// TIA Portal project "Respirator2020_V16" (V16)

(* hardware
DEVICE "S7-1200 station_1"  S7-1200 Station
   slot 0: "Rack_0"  S7-1200 Rack  Rack  V1.0
   slot 1: "PLC_1"  CPU 1215C DC/DC/DC  6ES7 215-1AG40-0XB0  V4.2
DEVICE "HMI_1"  TP700 Comfort
   slot 0: "HMI_1"  TP700 Comfort  6AV2 124-0GC01-0AX0  15.1.0.0
   slot 1: "HMI_RT_1"  TP700 Comfort  6AV2 124-0GC01-0AX0  15.1.0.0
   slot 5: "HMI_1.IE_CP_1"  PROFINET Interface  15.0.1.0
      slot 1: "Interfaz PROFINET_1"  PROFINET Interface
         slot 1: "Port_1"  Port
         slot 2: "Port_2"  Port
   slot 7: "HMI_1.MPI/DP_CP_1"  MPI/DP Interface  15.0.1.0
*)

// ===== PLC "PLC_1"  CPU 1215C DC/DC/DC =====

VAR_GLOBAL   // PLC tag table "Tabla de variables estándar"
   "System_Byte" AT %MB1 : Byte;
   "FirstScan" AT %M1.0 : Bool;
   "DiagStatusUpdate" AT %M1.1 : Bool;
   "AlwaysTRUE" AT %M1.2 : Bool;
   "AlwaysFALSE" AT %M1.3 : Bool;
   "Clock_Byte" AT %MB0 : Byte;
   "Clock_10Hz" AT %M0.0 : Bool;
   "Clock_5Hz" AT %M0.1 : Bool;
   "Clock_2.5Hz" AT %M0.2 : Bool;
   "Clock_2Hz" AT %M0.3 : Bool;
   "Clock_1.25Hz" AT %M0.4 : Bool;
   "Clock_1Hz" AT %M0.5 : Bool;
   "Clock_0.625Hz" AT %M0.6 : Bool;
   "Clock_0.5Hz" AT %M0.7 : Bool;
   "TurnAxisDir" AT %Q0.1 : Bool;
   "TurnAxisPulse" AT %Q0.0 : Bool;
   "EmergencyStop" AT %I0.0 : Bool;
   "ServoPend" AT %I1.0 : Bool;
   "ServoAlarm" AT %I1.1 : Bool;
   "TurnAxisEnable" AT %Q0.2 : Bool;
   "AtmosfericPressure" AT %IW64 : Int;
   "DiferentialPressure" AT %IW66 : Int;
   "TurnAxisHwLow" AT %I1.2 : Bool;
   "TurnAxisHwHi" AT %I1.3 : Bool;
   "HW_PWN_DutyCicle" AT %QW1008 : Hw_Pwm;
   "HW_PWM_Frecuency" AT %QD1010 : DInt;
   "COM_METEO_CONFIGURATION" AT %M202.0 : Bool;
   "COM_METEO_RESET" AT %M202.1 : Bool;
   "COM_METEO_DELETE_BUFFER" AT %M202.2 : Bool;
   "COM_METEO_RECEIVE" AT %M202.3 : Bool;
   "COM_METEO_SEND" AT %M202.4 : Bool;
   "COM_METEO_CHECKSUM" AT %M202.5 : Bool;
   "ResetComm" AT %M100.0 : Bool;
   "PeepValve" AT %Q0.4 : Bool;
   "Buzzer" AT %Q1.1 : Bool;
   "BeaconLightRed" AT %Q0.6 : Bool;
   "BeaconLightOrange" AT %Q0.7 : Bool;
   "BeaconLightGreen" AT %Q1.0 : Bool;
   "ResetRelay" AT %Q0.5 : Bool;
   "Tag_1" AT %M10.0 : Bool;
END_VAR

VAR_GLOBAL CONSTANT   // PLC tag table "Tabla de variables estándar"
   "Startup1" : Int := 1;
   "Configuration" : Int := 2;
   "Delete_Buffer" : Int := 3;
   "Data_Reception" : Int := 4;
   "Data_Transmision" : Int := 5;
   "STOP" : Int := 0;
END_VAR

TYPE "Motor"
   STRUCT
      POWER_ENABLE : Bool;
      POWER_START_MODE : Int;
      POWER_STOP_MODE : Int;
      POWER_STATUS : Bool;
      POWER_BUSY : Bool;
      POWER_ERROR : Bool;
      POWER_ERROR_ID : Int;
      POWER_ERROR_INFO : Int;
      RESET_EXECUTE : Bool;
      RESET_RESTART : Bool;
      RESET_DONE : Bool;
      RESET_BUSY : Bool;
      RESET_ERROR : Bool;
      RESET_ERROR_ID : Int;
      RESET_ERROR_INFO : Int;
      HOME_EXECUTE : Bool;
      HOME_POSITION : Real;
      HOME_MODE : Int;
      HOME_DONE : Bool;
      HOME_BUSY : Bool;
      HOME_COMMAND_ABORTED : Bool;
      HOME_ERROR : Bool;
      HOME_ERROR_ID : Int;
      HOME_ERROR_INFO : Int;
      HOME_REFERENCE_MARK_POS : Real;
      HALT_EXECUTE : Bool;
      HALT_DONE : Bool;
      HALT_BUSY : Bool;
      HALT_COMMAND_ABORTED : Bool;
      HALT_ERROR : Bool;
      HALT_ERROR_ID : Int;
      HALT_ERROR_INFO : Int;
      JOG_FORWARD : Bool;
      JOG_BACKWARD : Bool;
      JOG_VELOCITY : Real;
      JOG_POSITION_CONTROLLED : Bool;
      JOG_IN_VELOCITY : Bool;
      JOG_BUSY : Bool;
      JOG_COMMAND_ABORTED : Bool;
      JOG_ERROR : Bool;
      JOG_ERROR_ID : Int;
      JOG_ERROR_INFO : Int;
      ABSOLUTE_EXECUTE : Bool;
      ABSOLUTE_POSITION : Real;
      ABSOLUTE_VELOCITY : Real;
      ABSOLUTE_DIRECTION : Int;
      ABSOLUTE_DONE : Bool;
      ABSOLUTE_BUSY : Bool;
      ABSOLUTE_COMMAND_ABORTED : Bool;
      ABSOLUTE_ERROR : Bool;
      ABSOLUTE_ERROR_ID : Int;
      ABSOLUTE_ERROR_INFO : Int;
   END_STRUCT;
END_TYPE

TYPE "DTAlarm"
   STRUCT
      ENTERADO : Bool;
      REARME : Bool;
      FUNCION : Bool;
      ENTRADA : Bool;
      SALIDA_VISUALIZACION : Bool;
      SALIDA_VISUALIZACION_NEGADA : Bool;
      SALIDA_ENCLAVAMIENTO : Bool;
      SALIDA_ENCLAVAMIENTO_NEGADA : Bool;
   END_STRUCT;
END_TYPE

TYPE "DTAlarmSPV"
   STRUCT
      ENTERADO : Bool;
      REARME : Bool;
      FUNCION : Int;
      ENTRADA_ALM : Bool;
      ENTRADA_SPV : Bool;
      ORDEN_MARCHA : Bool;
      RETARDO : Time;
      SALIDA_VISUALIZACION : Bool;
      SALIDA_VISUALIZACION_NEGADA : Bool;
      SALIDA_ENCLAVAMIENTO : Bool;
      SALIDA_ENCLAVAMIENTO_NEGADA : Bool;
      SALIDA_SUPERVISION : Bool;
      T_TRANSCURRIDO : Time;
   END_STRUCT;
END_TYPE

// folder: 1_Data

DATA_BLOCK "Data_DB"   // DB10
{ S7_Optimized_Access := 'TRUE' }
AUTHOR : JL_Cristobal_2020
VERSION : 0.1
// stored: InstanceOfName Data
"Data"
BEGIN
END_DATA_BLOCK

DATA_BLOCK "TidalVolumeCalculator_DB"   // DB11
{ S7_Optimized_Access := 'TRUE' }
AUTHOR : JL_Cristobal_2020
VERSION : 0.1
// stored: InstanceOfName TidalVolumeCalculator
"TidalVolumeCalculator"
BEGIN
END_DATA_BLOCK

DATA_BLOCK "DataValues"   // DB101
{ S7_Optimized_Access := 'TRUE' }
AUTHOR : JL_Cristobal_2020
VERSION : 0.1
   VAR
      FlowRaw : Real;
      FlowValue : Real;
      DiferntialPressureRaw : Real;
      DiferntialPressure : Real;
      PipValue : Real;
      PlateauValue : Real;
      PeepValue : Real;
      FrequencyValue : Real;
      TidalVolumeValue : Real;
      VolumeMinuteValue : Real;
      Trigger : Real;
      DrivingPressure : Real;
      BatteryVoltage : Real;
      BatteryCapacity : Real;
      Pressure1 : Real;
      Pressure2 : Real;
      VomumeAccumulated : Real;
      Flow : Real;
      AirPressure : Real;
      O2Pressure : Real;
      CalculatedRatio : Real;
      InspirationTime : Time;
      RestTime : Time;
      EspirationTime : Time;
      DelayTime : Time;
      TotalTime : Time;
   END_VAR
BEGIN
END_DATA_BLOCK

DATA_BLOCK "DateTime"   // DB102
{ S7_Optimized_Access := 'FALSE' }
AUTHOR : JL_Cristobal_2020
VERSION : 0.1
   VAR
      SystemDateRetVal : Int;
      SystemDateOut : DTL;
      LocalDateRetVal : Int;
      LocalDateOut : DTL;
      WriteDateTime : DTL;
      WriteDateOut : Int;
      SetWriteData : Bool;
      StatuSetTime : DTL;
      SetTime : Bool;
      INT_FS : DWord;
      INT_FC : DWord;
      INT_HS : DWord;
      INT_HC : DWord;
      SystemDate_W : Word;
      SystemTime_W : Word;
   END_VAR
BEGIN
END_DATA_BLOCK

DATA_BLOCK "OperatingParameters"   // DB103
{ S7_Optimized_Access := 'TRUE' }
AUTHOR : JL_Cristobal_2020
VERSION : 0.1
   VAR RETAIN
      PipMax : Real := 40.0;
      PipSetpoint : Real := 20.0;
      PipMin : Real := 10.0;
      PipFactor : Real := 1.0;
      PlateauMax : Real;
      PlateauSetpoint : Real;
      PlateauMin : Real;
      PlateauFactor : Real := 1.0;
      PeepMax : Real := 15.0;
      PeepSetpoint : Real := 8.0;
      PeepMin : Real := 6.0;
      PeepFactor : Real;
      FrequencyMax : Real := 24.0;
      FrequencySetpoint : Real := 10.0;
      FrequencyMin : Real := 3.0;
      FrequencyFactor : Real := 1.0;
      TidalVolumenMax : Real := 900.0;
      TidalVolumenSetpoint : Real := 400.0;
      TidalVolumenMin : Real := 100.0;
      TidalVolumenFactor : Real := 1.0;
      VolumeMinMax : Real;
      VolumeMinSetpoint : Real;
      VolumeMinMin : Real;
      VolumeMinFactor : Real := 1.0;
      TriggerMax : Real;
      TriggerSetpoint : Real := 10.0;
      TriggerMin : Real;
      TriggerFactor : Real := 1.0;
      Trigger : Bool;
      AirMax : Real;
      AirSetpoint : Real := 10.0;
      AirMin : Real;
      AirFactor : Real := 1.0;
      Air : Bool;
      O2Max : Real;
      O2Setpoint : Real := 10.0;
      O2Min : Real;
      O2Factor : Real := 1.0;
      O2 : Bool;
      InpirationRatio : Real;
      EspirationRatio : Real;
      DelayRatio : Real;
   END_VAR
   VAR
      RestRatio : Real;
      CalculatedRatio : Real;
   END_VAR
   VAR RETAIN
      BatteryLevelTrigger : Real := 22.0;
   END_VAR
   VAR
      PeakPBPlus : Bool;
      PeakPBMinus : Bool;
      PeepPBPlus : Bool;
      PeepPBMinus : Bool;
      FrPBPlus : Bool;
      FrPBMinus : Bool;
      RecruitmentOn : Bool;
      RecruitmentOff : Bool;
      RecruitmentMem : Bool;
      RecruitmentRunning : Bool;
      RecruitmentEnding : Bool;
      RecruitmentEnd : Bool;
   END_VAR
   VAR RETAIN
      RecruitmentTimer : Time := T#40s;
   END_VAR
   VAR
      RecruitmentElap : Time;
   END_VAR
   VAR RETAIN
      HumidifierTimer : Time := T#40s;
   END_VAR
   VAR
      HumidifiertElap : Time;
   END_VAR
   VAR RETAIN
      HumidifiertDuration : Time;
      ControlMode : Int;
   END_VAR
BEGIN
END_DATA_BLOCK

DATA_BLOCK "PatientData"   // DB104
{ S7_Optimized_Access := 'TRUE' }
AUTHOR : JL_Cristobal_2020
VERSION : 0.1
   VAR RETAIN
      PatientType : Int;
      PatientWeight : Real;
      PatientHeight : Real;
   END_VAR
   VAR
      TidalVolume : Real;
   END_VAR
   VAR RETAIN
      TimeStart : Time_Of_Day;
      TimeEnd : Time_Of_Day;
   END_VAR
BEGIN
END_DATA_BLOCK

DATA_BLOCK "ProcessData"   // DB105
{ S7_Optimized_Access := 'TRUE' }
NAME : JL_Cristobal_2020
VERSION : 0.1
   VAR
      PIDSetpoint : Real;
      PIDErrorAck : Bool;
      PIDInput : Real;
      PIDInput_PER : Int;
      PIDReset : Bool;
      PIDModeActivate : Bool;
      PIDMode : Int;
      PIDInterlock : Bool;
      PIDOutReal : Real;
      PIDOutInt : Int;
      PIDOutPWM : Bool;
      PIDState : Int;
      PIDError : Bool;
      PIDErrorBits : Int;
      PIDOutMotor : Real;
   END_VAR
   VAR RETAIN
      PipSetpointPreAlarmHI : Real;
      PpipSetpointAlarmHI : Real;
      PipSetpointPreAlarmLOW : Real;
      PipSetpointAlarmLOW : Real;
      PipSetpointHysteresisHI : Real;
      PipSetpointHysteresisLOW : Real;
      PlateauSetpointPreAlarmHI : Real;
      PlateauSetpointAlarmHI : Real;
      PlateauSetpointPreAlarmLOW : Real;
      PlateauSetpointAlarmLOW : Real;
      PlateauSetpointHysteresisHI : Real;
      PlateauSetpointHysteresisLOW : Real;
      PeepSetpointPreAlarmHI : Real;
      PeepSetpointAlarmHI : Real;
      PeepSetpointPreAlarmLOW : Real;
      PeepSetpointAlarmLOW : Real;
      PeepSetpointHysteresisHI : Real;
      PeepSetpointHysteresisLOW : Real;
      FrequencySetpointPreAlarmHI : Real;
      FrequencySetpointAlarmHI : Real;
      FrequencySetpointPreAlarmLOW : Real;
      FrequencySetpointAlarmLOW : Real;
      FrequencySetpointHysteresisHI : Real;
      FrequencySetpointHysteresisLOW : Real;
      TidalVolumeSetpointPreAlarmHI : Real;
      TidalVolumeSetpointAlarmHI : Real;
      TidalVolumeSetpointPreAlarmLOW : Real;
      TidalVolumeSetpointAlarmLOW : Real;
      TidalVolumeHystersisHI : Real;
      TidalVolumeHystersisLOW : Real;
      VolumeMinSetpointPreAlarmHI : Real;
      VolumeMinSetpointAlarmHI : Real;
      VolumeMinSetpointPreAlarmLOW : Real;
      VolumeMinSetpointAlarmLOW : Real;
      VolumeMinHysteresisHI : Real;
      VolumeMinHysteresisLOW : Real;
      TriggeVolumeSetpointPreAlarmHI : Real;
      TriggerVolumeSetpointAlarmHI : Real;
      TriggerVolumeSetpointPreAlarmLOW : Real;
      TriggerVolumeSetpointAlarmLOW : Real;
      TriggerVolumeHysteresisHI : Real;
      TriggerVolumeHysteresisLOW : Real;
      BatterySetpointPreAlarmHI : Real := 27.0;
      BatterySetpointAlarmHI : Real := 26.0;
      BatterySetpointPreAlarmLOW : Real := 23.0;
      BatterySetpointAlarmLOW : Real := 22.0;
      BatterySetpointHysteresisHI : Real;
      BatterySetpointHysteresisLOW : Real;
      AirSetpointPreAlarmHI : Real := 27.0;
      AirSetpointAlarmHI : Real := 26.0;
      AirSetpointPreAlarmLOW : Real := 23.0;
      AirSetpointAlarmLOW : Real := 22.0;
      AirSetpointHysteresisHI : Real;
      AirSetpointHysteresisLOW : Real;
      O2SetpointPreAlarmHI : Real := 27.0;
      O2SetpointAlarmHI : Real := 26.0;
      O2SetpointPreAlarmLOW : Real := 23.0;
      "02SetpointAlarmLOW" : Real := 22.0;
      O2SetpointHysteresisHI : Real;
      O2SetpointHysteresisLOW : Real;
   END_VAR
BEGIN
END_DATA_BLOCK

DATA_BLOCK "RatioCalculator_DB"   // DB106
{ S7_Optimized_Access := 'TRUE' }
AUTHOR : JL_Cristobal_2020
VERSION : 0.1
// stored: InstanceOfName RatioCalculator
"RatioCalculator"
BEGIN
END_DATA_BLOCK

DATA_BLOCK "VariableSupervisor_DB_Frecuency"   // DB120
{ S7_Optimized_Access := 'TRUE' }
AUTHOR : JL_Cristobal_2020
VERSION : 0.1
// stored: InstanceOfName VariableSupervisor
"VariableSupervisor"
BEGIN
END_DATA_BLOCK

DATA_BLOCK "VariableSupervisor_DB_Peep"   // DB121
{ S7_Optimized_Access := 'TRUE' }
AUTHOR : JL_Cristobal_2020
VERSION : 0.1
// stored: InstanceOfName VariableSupervisor
"VariableSupervisor"
BEGIN
END_DATA_BLOCK

DATA_BLOCK "VariableSupervisor_DB_Pip"   // DB122
{ S7_Optimized_Access := 'TRUE' }
AUTHOR : JL_Cristobal_2020
VERSION : 0.1
// stored: InstanceOfName VariableSupervisor
"VariableSupervisor"
BEGIN
END_DATA_BLOCK

DATA_BLOCK "VariableSupervisor_DB_Plateau"   // DB123
{ S7_Optimized_Access := 'TRUE' }
AUTHOR : JL_Cristobal_2020
VERSION : 0.1
// stored: InstanceOfName VariableSupervisor
"VariableSupervisor"
BEGIN
END_DATA_BLOCK

DATA_BLOCK "VariableSupervisor_DB_TidalVolume"   // DB124
{ S7_Optimized_Access := 'TRUE' }
AUTHOR : JL_Cristobal_2020
VERSION : 0.1
// stored: InstanceOfName VariableSupervisor
"VariableSupervisor"
BEGIN
END_DATA_BLOCK

DATA_BLOCK "VariableSupervisor_DB_Trigger"   // DB125
{ S7_Optimized_Access := 'TRUE' }
AUTHOR : JL_Cristobal_2020
VERSION : 0.1
// stored: InstanceOfName VariableSupervisor
"VariableSupervisor"
BEGIN
END_DATA_BLOCK

DATA_BLOCK "VariableSupervisor_DB_VolumeMin"   // DB126
{ S7_Optimized_Access := 'TRUE' }
AUTHOR : JL_Cristobal_2020
VERSION : 0.1
// stored: InstanceOfName VariableSupervisor
"VariableSupervisor"
BEGIN
END_DATA_BLOCK

// folder: 2_SensorComm

DATA_BLOCK "SensorComm_PtP_Freeport_DB"   // DB20
{ S7_Optimized_Access := 'FALSE' }
AUTHOR : JL_Cristobal_2020
VERSION : 0.1
// stored: InstanceOfName SensorComm_PtP_Freeport
"SensorComm_PtP_Freeport"
BEGIN
END_DATA_BLOCK

DATA_BLOCK "SensorComm_A_Port_Config_Settings"   // DB200
{ S7_Optimized_Access := 'FALSE' }
AUTHOR : JL_Cristobal_2020
VERSION : 0.1
   VAR
      Protocol : Word := 16#0000;
      Baud : Word := 16#0009;
      Parity : Word := 16#0001;
      DataBits : Word := 16#0001;
      StopBits : Word := 16#0001;
      FLOWCTRL : Word := 16#0001;
      XonChar : Char := ' ';
      XoffChar : Char := ' ';
      WaitTime : Word := 16#0000;
      Mode : Byte := 16#00;
      LinePre : Byte := 16#00;
      BrkDet : Byte;
      UserInt : Bool := FALSE;
      Output : Struct
         Done : Bool := FALSE;
         Error : Bool := FALSE;
         Status : DWord := 16#0000_0000;
         State : Int := 2;
         RingPlace : Int := 0;
         Lenght : Int := 0;
      END_STRUCT;
   END_VAR
BEGIN
END_DATA_BLOCK

DATA_BLOCK "SensorComm_B_PtP_Freeport_DB"   // DB201
{ S7_Optimized_Access := 'FALSE' }
AUTHOR : JL_Cristobal_2020
VERSION : 0.1
// stored: InstanceOfName SensorComm_PtP_Freeport
"SensorComm_PtP_Freeport"
BEGIN
END_DATA_BLOCK

DATA_BLOCK "SensorComm_C_buffer_ptp"   // DB202
{ S7_Optimized_Access := 'FALSE' }
AUTHOR : JL_Cristobal_2020
VERSION : 0.1
   VAR
      Ringbuffer : Array[0..1024] of Char;
   END_VAR
BEGIN
END_DATA_BLOCK

DATA_BLOCK "SensorComm_D_Commands"   // DB203
{ S7_Optimized_Access := 'TRUE' }
AUTHOR : JL_Cristobal_2020
VERSION : 0.1
   VAR RETAIN
      Commands : Struct
         Command1 : String := 'M9';
         Command2 : String := 'Co';
         Command3 : String := 'IN';
         Command4 : String := 'CA';
         Command5 : String := 'NE';
         Command6 : String := 'FA';
         Command7 : String := 'AI';
         Command8 : String := 'S\';
         Command9 : String := 'M\';
         Command10 : String := 'D\';
         Command11 : String := 'T1';
         Command12 : String;
      END_STRUCT;
   END_VAR
BEGIN
END_DATA_BLOCK

DATA_BLOCK "SensorComm_E_Data"   // DB204
{ S7_Optimized_Access := 'TRUE' }
AUTHOR : JL_Cristobal_2020
VERSION : 0.1
   VAR
      Read : String;
      OpretingMode : Int;
      OutputStatus : Struct
         Pressure1 : Real;
         Pressure2 : Real;
         VolumeAccumulated : Real;
         Flow : Real;
         ErrorPressure1 : Bool;
         ErrorPressure2 : Bool;
         ErrorVolumeAccumulated : Bool;
         ErrorFlux : Bool;
      END_STRUCT;
   END_VAR
BEGIN
END_DATA_BLOCK

// folder: 3_Alarms

DATA_BLOCK "Alarm0Pack16B"   // DB300
{ S7_Optimized_Access := 'FALSE' }
AUTHOR : JL_Cristobal_2020
VERSION : 0.1
// stored: InstanceOfName Pack_16B
"Pack_16B"
BEGIN
END_DATA_BLOCK

DATA_BLOCK "Alarm1Pack16B"   // DB301
{ S7_Optimized_Access := 'FALSE' }
AUTHOR : JL_Cristobal_2020
VERSION : 0.1
// stored: InstanceOfName Pack_16B
"Pack_16B"
BEGIN
END_DATA_BLOCK

DATA_BLOCK "Alarm2Pack16B"   // DB302
{ S7_Optimized_Access := 'FALSE' }
AUTHOR : JL_Cristobal_2020
VERSION : 0.1
// stored: InstanceOfName Pack_16B
"Pack_16B"
BEGIN
END_DATA_BLOCK

DATA_BLOCK "Alarm3Pack16B"   // DB303
{ S7_Optimized_Access := 'FALSE' }
AUTHOR : JL_Cristobal_2020
VERSION : 0.1
// stored: InstanceOfName Pack_16B
"Pack_16B"
BEGIN
END_DATA_BLOCK

DATA_BLOCK "AlarmsCall_DB"   // DB304
{ S7_Optimized_Access := 'TRUE' }
AUTHOR : JL_Cristobal_2020
VERSION : 0.1
// stored: InstanceOfName Alarms
"Alarms"
BEGIN
END_DATA_BLOCK

DATA_BLOCK "AlarmsRaw"   // DB305
{ S7_Optimized_Access := 'TRUE' }
AUTHOR : JL_Cristobal_2020
VERSION : 0.1
   VAR
      PipDisplayPreAlarmHI : Bool;
      PipDisplayAlarmHI : Bool;
      PipDisplayPreAlarmLOW : Bool;
      PipDisplayAlarmLOW : Bool;
      PipInterlockPreAlarmHI : Bool;
      PipInterlockAlarmHI : Bool;
      PipInterlockPreAlarmLOW : Bool;
      PipInterlockAlarmLOW : Bool;
      PlateauDisplayPreAlarmHI : Bool;
      PlateauDisplayAlarmHI : Bool;
      PlateauDisplayPreAlarmLOW : Bool;
      PlateauDisplayAlarmLOW : Bool;
      PlateauInterlockPreAlarmHI : Bool;
      PlateauInterlockAlarmHI : Bool;
      PlateauInterlockPreAlarmLOW : Bool;
      PlateauInterlockAlarmLOW : Bool;
      PeepDisplayPreAlarmHI : Bool;
      PeepDisplayAlarmHI : Bool;
      PeepDisplayPreAlarmLOW : Bool;
      PeepDisplayAlarmLOW : Bool;
      PeepInterlockPreAlarmHI : Bool;
      PeepInterlockAlarmHI : Bool;
      PeepInterlockPreAlarmLOW : Bool;
      PeepInterlockAlarmLOW : Bool;
      FrequencyDisplayPreAlarmHI : Bool;
      FrequencyDisplayAlarmHI : Bool;
      FrequencyDisplayPreAlarmLOW : Bool;
      FrequencyDisplayAlarmLOW : Bool;
      FrequencyInterlockPreAlarmHI : Bool;
      FrequencyInterlockAlarmHI : Bool;
      FrequencyInterlockPreAlarmLOW : Bool;
      FrequencyInterlockAlarmLOW : Bool;
      TidalVolumeDisplayPreAlarmHI : Bool;
      TidalVolumeDisplayAlarmHI : Bool;
      TidalVolumeDisplayPreAlarmLOW : Bool;
      TidalVolumeDisplayAlarmLOW : Bool;
      TidalVolumeInterlockPreAlarmHI : Bool;
      TidalVolumeInterlockAlarmHI : Bool;
      TidalVolumeInterlockPreAlarmLOW : Bool;
      TidalVolumeInterlockAlarmLOW : Bool;
      VolumeMinuteDisplayPreAlarmHI : Bool;
      VolumeMinuteDisplayAlarmHI : Bool;
      VolumeMinuteDisplayPreAlarmLOW : Bool;
      VolumeMinuteDisplayAlarmLOW : Bool;
      VolumeMinuteInterlockPreAlarmHI : Bool;
      VolumeMinuteInterlockAlarmHI : Bool;
      VolumeMinuteInterlockPreAlarmLOW : Bool;
      VolumeMinuteInterlockAlarmLOW : Bool;
      TriggerDisplayPreAlarmHI : Bool;
      TriggerDisplayAlarmHI : Bool;
      TriggerDisplayPreAlarmLOW : Bool;
      TriggerDisplayAlarmLOW : Bool;
      TriggerInterlockPreAlarmHI : Bool;
      TriggerInterlockAlarmHI : Bool;
      TriggerInterlockPreAlarmLOW : Bool;
      TriggerInterlockAlarmLOW : Bool;
      BatteryDisplayPreAlarmHI : Bool;
      BatteryDisplayAlarmHI : Bool;
      BatteryDisplayPreAlarmLOW : Bool;
      BatteryDisplayAlarmLOW : Bool;
      BatteryInterlockPreAlarmHI : Bool;
      BatteryInterlockAlarmHI : Bool;
      BatteryInterlockPreAlarmLOW : Bool;
      BatteryInterlockAlarmLOW : Bool;
   END_VAR
BEGIN
END_DATA_BLOCK

DATA_BLOCK "AlarmsWord"   // DB306
{ S7_Optimized_Access := 'FALSE' }
AUTHOR : JL_Cristobal_2020
VERSION : 0.1
   VAR
      Alarms : Array[0..100] of Word;
   END_VAR
BEGIN
   Alarms[0] := 0;
END_DATA_BLOCK

DATA_BLOCK "DirectAnalog_DB_Battery"   // DB310
{ S7_Optimized_Access := 'FALSE' }
AUTHOR : JL_Cristobal_2020
VERSION : 0.1
// stored: InstanceOfName DirectAnalog
"DirectAnalog"
BEGIN
END_DATA_BLOCK

DATA_BLOCK "DirectAnalog_DB_Frequency"   // DB311
{ S7_Optimized_Access := 'FALSE' }
AUTHOR : JL_Cristobal_2020
VERSION : 0.1
// stored: InstanceOfName DirectAnalog
"DirectAnalog"
BEGIN
END_DATA_BLOCK

DATA_BLOCK "DirectAnalog_DB_Peak"   // DB312
{ S7_Optimized_Access := 'FALSE' }
AUTHOR : JL_Cristobal_2020
VERSION : 0.1
// stored: InstanceOfName DirectAnalog
"DirectAnalog"
BEGIN
END_DATA_BLOCK

DATA_BLOCK "DirectAnalog_DB_Peep"   // DB313
{ S7_Optimized_Access := 'FALSE' }
AUTHOR : JL_Cristobal_2020
VERSION : 0.1
// stored: InstanceOfName DirectAnalog
"DirectAnalog"
BEGIN
END_DATA_BLOCK

DATA_BLOCK "DirectAnalog_DB_Plateau"   // DB314
{ S7_Optimized_Access := 'FALSE' }
AUTHOR : JL_Cristobal_2020
VERSION : 0.1
// stored: InstanceOfName DirectAnalog
"DirectAnalog"
BEGIN
END_DATA_BLOCK

DATA_BLOCK "DirectAnalog_DB_TidalVolume"   // DB315
{ S7_Optimized_Access := 'FALSE' }
AUTHOR : JL_Cristobal_2020
VERSION : 0.1
// stored: InstanceOfName DirectAnalog
"DirectAnalog"
BEGIN
END_DATA_BLOCK

DATA_BLOCK "DirectAnalog_DB_Trigger"   // DB316
{ S7_Optimized_Access := 'FALSE' }
AUTHOR : JL_Cristobal_2020
VERSION : 0.1
// stored: InstanceOfName DirectAnalog
"DirectAnalog"
BEGIN
END_DATA_BLOCK

DATA_BLOCK "DirectAnalog_DB_VolumeMinute"   // DB317
{ S7_Optimized_Access := 'FALSE' }
AUTHOR : JL_Cristobal_2020
VERSION : 0.1
// stored: InstanceOfName DirectAnalog
"DirectAnalog"
BEGIN
END_DATA_BLOCK

// folder: 4_ProcessControl

DATA_BLOCK "kkl_DB"   // DB15
{ S7_Optimized_Access := 'TRUE' }
AUTHOR : JL_Cristobal_2020
VERSION : 0.1
// stored: InstanceOfName 0_ProcessControl
"0_ProcessControl"
BEGIN
END_DATA_BLOCK

DATA_BLOCK "0_ProcessControl_DB"   // DB40
{ S7_Optimized_Access := 'TRUE' }
AUTHOR : JL_Cristobal_2020
VERSION : 0.1
// stored: InstanceOfName 0_ProcessControl
"0_ProcessControl"
BEGIN
END_DATA_BLOCK

DATA_BLOCK "2_PWMValve"   // DB400
{ S7_Optimized_Access := 'TRUE' }
AUTHOR : JL_Cristobal_2020
VERSION : 0.1
   VAR
      Enable : Bool;
      Busy : Bool;
      Status : Int;
      Frecuency : DInt;
      Duty_Cycle : Int;
   END_VAR
BEGIN
END_DATA_BLOCK

DATA_BLOCK "MotorControl"   // DB401
{ S7_Optimized_Access := 'TRUE' }
AUTHOR : JL_Cristobal_2020
VERSION : 0.1
   VAR
      POWER_Enable : Bool;
      POWER_StartMode : Int;
      POWER_StopMode : Int;
      POWER_Status : Bool;
      POWER_Error : Bool;
      ReadyMotor : Bool;
      RESET_Execute : Bool;
      RESET_Done : Bool;
      RESET_Error : Bool;
      HOME_Execute : Bool;
      HOME_Position : Real;
   END_VAR
   VAR RETAIN
      HOME_Mode : Int := 3;
   END_VAR
   VAR
      HOME_Done : Bool;
      HOME_Error : Bool;
      HALT_Execute : Bool;
      HALT_Done : Bool;
      HALT_Error : Bool;
      ABSOLUTE_Execute : Bool;
      ABSOLUTE_Position : Real;
      ABSOLUTE_Velocity : Real;
      ABSOLUTE_Done : Bool;
      ABSOLUTE_Error : Bool;
      RELATIVE_Execute : Bool;
      RELATIVE_Distance : Real;
      RELATIVE_Velocity : Real;
      RELATIVE_Done : Bool;
      RELATIVE_Error : Bool;
      Velocity_Execute : Bool;
      Velocity_Velocity : Real;
      Velocity_Current : Bool;
      Velocity_invelocity : Bool;
      Velocity_Error : Bool;
      JOG_Forward : Bool;
      JOG_Backward : Bool;
      JOG_Velocity : Real;
      JOG_Invelocity : Bool;
      JOG_Error : Bool;
      Permissions : Bool;
   END_VAR
BEGIN
END_DATA_BLOCK

DATA_BLOCK "Operation"   // DB402
{ S7_Optimized_Access := 'TRUE' }
AUTHOR : JL_Cristobal_2020
VERSION : 0.1
   VAR
      Operation_ON : Bool;
      Emergency : Bool;
      GeneralAck : Bool;
      MotorAck : Bool;
      ProcessAck : Bool;
      GeneralReset : Bool;
      MotorReset : Bool;
      ProcessReset : Bool;
      LampTest : Bool;
      RecruimentSignal : Bool;
      RecruimentSignalEnding : Bool;
      InterlockPip : Bool;
      InterlockPlateau : Bool;
      InterlockPeep : Bool;
      InterlockFrequency : Bool;
      InterlockTidalVomume : Bool;
      InterlockVolMinute : Bool;
      InterlockTrigger : Bool;
      InterlockBattery : Bool;
   END_VAR
BEGIN
END_DATA_BLOCK

DATA_BLOCK "PIDData"   // DB403
{ S7_Optimized_Access := 'TRUE' }
AUTHOR : JL_Cristobal_2020
VERSION : 0.1
   VAR
      A_Setpoint : Real;
      A_Input : Real;
      A_InputPER : Real;
      A_ErrorACK : Bool;
      A_Reset : Bool;
      A_ModeActivate : Bool;
      A_Mode : Int;
      A_Interlock : Bool;
      B_Setpoint : Real;
      B_Input : Real;
      B_InputPER : Real;
      B_ErrorACK : Bool;
      B_Reset : Bool;
      B_ModeActivate : Bool;
      B_Mode : Int;
      B_Interlock : Bool;
      C_Setpoint : Real;
      C_Input : Real;
      C_InputPER : Real;
      C_ErrorACK : Bool;
      C_Reset : Bool;
      C_ModeActivate : Bool;
      C_Mode : Int;
      C_Interlock : Bool;
      D_Setpoint : Real;
      D_Input : Real;
      D_InputPER : Real;
      D_ErrorACK : Bool;
      D_Reset : Bool;
      D_ModeActivate : Bool;
      D_Mode : Int;
      D_Interlock : Bool;
      ChannelSelect : Int;
   END_VAR
BEGIN
END_DATA_BLOCK

DATA_BLOCK "PIDSwitch_DB"   // DB404
{ S7_Optimized_Access := 'TRUE' }
AUTHOR : JL_Cristobal_2020
VERSION : 0.1
// stored: InstanceOfName PIDSwitch
"PIDSwitch"
BEGIN
END_DATA_BLOCK

// folder: System blocks/Program resources

DATA_BLOCK "IEC_Timer_0_DB_SPV"   // DB33
{ S7_Optimized_Access := 'TRUE' }
AUTHOR : Simatic
FAMILY : IEC
NAME : IEC_TMR
VERSION : 1.0
// stored: InstanceOfName IEC_TIMER
"IEC_TIMER"
BEGIN
END_DATA_BLOCK

DATA_BLOCK "IEC_Timer_0_DB_Recruitment"   // DB45
{ S7_Optimized_Access := 'TRUE' }
AUTHOR : Simatic
FAMILY : IEC
NAME : IEC_TMR
VERSION : 1.0
// stored: InstanceOfName IEC_TIMER
"IEC_TIMER"
BEGIN
END_DATA_BLOCK

DATA_BLOCK "IEC_Timer_0_DB_MotorEnable"   // DB50
{ S7_Optimized_Access := 'TRUE' }
AUTHOR : Simatic
FAMILY : IEC
NAME : IEC_TMR
VERSION : 1.0
// stored: InstanceOfName IEC_TIMER
"IEC_TIMER"
BEGIN
END_DATA_BLOCK

DATA_BLOCK "IEC_Timer_0_DB_Reset"   // DB51
{ S7_Optimized_Access := 'TRUE' }
AUTHOR : Simatic
FAMILY : IEC
NAME : IEC_TMR
VERSION : 1.0
// stored: InstanceOfName IEC_TIMER
"IEC_TIMER"
BEGIN
END_DATA_BLOCK

// folder: (top level)

DATA_BLOCK "TurnAxis"   // DB1, Motion_DB
{ S7_Optimized_Access := 'TRUE' }
AUTHOR : SIMATIC
FAMILY : BasicMC
NAME : TO_PosAx
VERSION : 6.0
// stored: InstanceOfName TO_PositioningAxis
"TO_PositioningAxis"
BEGIN
   // Axis.PositionLimitsMax_AddressCU = %I1.3
   // Axis.HomingReferencePointSwitch_AddressCU = %I1.2
   // Axis.PassiveHomingReferencePointSwitch_AddressCU = %I1.2
   // Axis.PositionLimitsMin_AddressCU = %I1.2
   // Axis.DirectionOutputEnabledCU = TRUE
   // Axis.OnlinePtoModeCU = 16#0000_0002
   // Axis.SelectedChannel2EnumCU = %Q0.1
   // Axis.SelectedChannel1EnumCU = %Q0.0
   // Pulse.MinDeltaDeltaFrequencyCU = 0.004
   // Pulse.MaxDeltaDeltaFrequencyCU = 1.0E+10
   // Pulse.MinDeltaFrequencyCU = 0.005
   // Pulse.MaxDeltaFrequencyCU = 9.5E+9
   // Pulse.MinFrequencyCU = 1.0
   // Pulse.MaxFrequencyCU = 100000.0
   // Pulse.OutputSourceCU = 16#0000_0000
   // Axis.SelectPTO = 0
   // Axis.LengthUnit.LastDistance = 1005
END_DATA_BLOCK

ORGANIZATION_BLOCK "Main"   // OB1, LAD, ProgramCycle
TITLE = "Main Program Sweep (Cycle)"
{ S7_Optimized_Access := 'TRUE' }
AUTHOR : JL_Cristobal_2020
VERSION : 0.1
   VAR_INPUT
      Initial_Call : Bool;   // Initial call of this OB
      Remanence : Bool;   // =True, if remanent data are available
   END_VAR
BEGIN

REGION Network 1: Function Call Sensors Communications
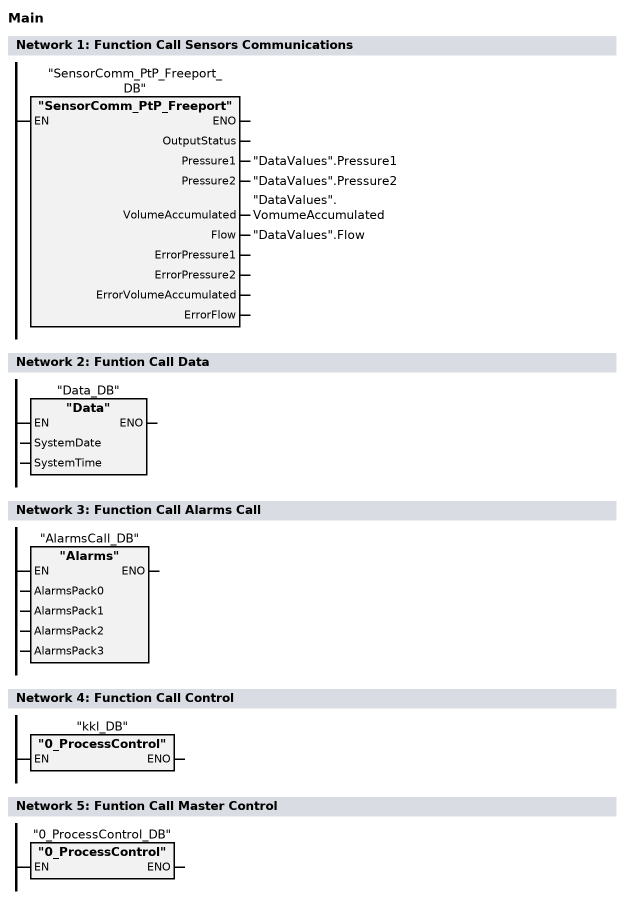
   RUNG wire#powerrail
      "SensorComm_PtP_Freeport_DB"(OutputStatus =>, Pressure1 => "DataValues".Pressure1, Pressure2 => "DataValues".Pressure2, VolumeAccumulated => "DataValues".VomumeAccumulated, Flow => "DataValues".Flow, ErrorPressure1 =>, ErrorPressure2 =>, ErrorVolumeAccumulated =>, ErrorFlow =>)
   END_RUNG
   // the same network as SCL:
   "SensorComm_PtP_Freeport_DB"(Pressure1 => "DataValues".Pressure1,   // "SensorComm_PtP_Freeport"
                           Pressure2 => "DataValues".Pressure2,
                           VolumeAccumulated => "DataValues".VomumeAccumulated,
                           Flow => "DataValues".Flow);
END_REGION

REGION Network 2: Funtion Call Data
   RUNG wire#powerrail
      "Data_DB"(SystemDate :=, SystemTime :=)
   END_RUNG
   // the same network as SCL:
   "Data_DB"();   // "Data"
END_REGION

REGION Network 3: Function Call Alarms Call
   RUNG wire#powerrail
      "AlarmsCall_DB"(AlarmsPack0 :=, AlarmsPack1 :=, AlarmsPack2 :=, AlarmsPack3 :=)
   END_RUNG
   // the same network as SCL:
   "AlarmsCall_DB"();   // "Alarms"
END_REGION

REGION Network 4: Function Call Control
   RUNG wire#powerrail
      "kkl_DB"()
   END_RUNG
   // the same network as SCL:
   "kkl_DB"();   // "0_ProcessControl"
END_REGION

REGION Network 5: Funtion Call Master Control
   RUNG wire#powerrail
      "0_ProcessControl_DB"()
   END_RUNG
   // the same network as SCL:
   "0_ProcessControl_DB"();   // "0_ProcessControl"
END_REGION
END_ORGANIZATION_BLOCK

ORGANIZATION_BLOCK "Cyclic interrupt_PID"   // OB30, LAD, CyclicInterrupt
{ S7_Optimized_Access := 'TRUE' }
AUTHOR : JL_Cristobal_2020
VERSION : 0.1
   VAR_INPUT
      Initial_Call : Bool;   // Initial call of this OB
      Event_Count : Int;   // Events discarded
   END_VAR
BEGIN

REGION Network 1: Flow Meter
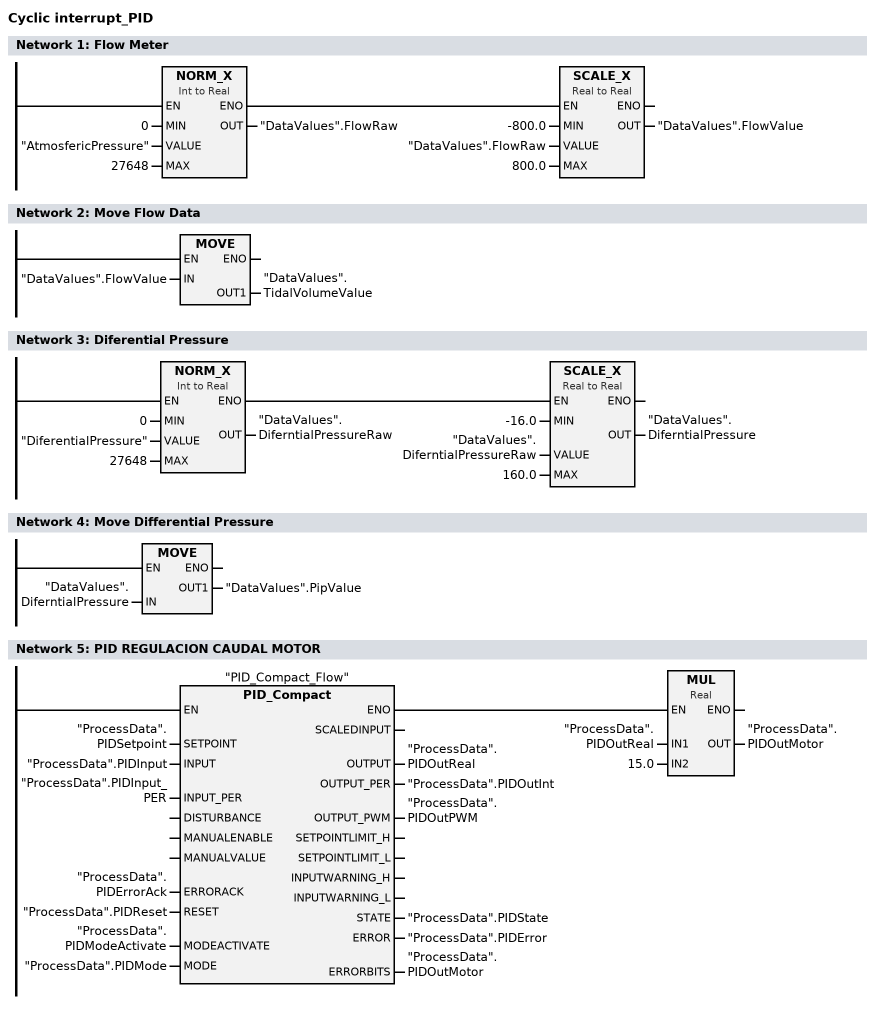
   RUNG wire#powerrail
      { S7_Templates := "[SrcType := Int, DestType := Real]" } Normalize(min := 0, value := "AtmosfericPressure", max := 27648, out => "DataValues".FlowRaw)
      { S7_Templates := "[SrcType := Real, DestType := Real]" } Scale(min := -800.0, value := "DataValues".FlowRaw, max := 800.0, out => "DataValues".FlowValue)
   END_RUNG
   // the same network as SCL:
   "DataValues".FlowRaw := NORM_X(MIN := 0, VALUE := "AtmosfericPressure", MAX := 27648);
   "DataValues".FlowValue := SCALE_X(MIN := -800.0, VALUE := "DataValues".FlowRaw, MAX := 800.0);
END_REGION

REGION Network 2: Move Flow Data
   RUNG wire#powerrail
      Move(in := "DataValues".FlowValue, out1 => "DataValues".TidalVolumeValue)
   END_RUNG
   // the same network as SCL:
   "DataValues".TidalVolumeValue := "DataValues".FlowValue;
END_REGION

REGION Network 3: Diferential Pressure
   RUNG wire#powerrail
      { S7_Templates := "[SrcType := Int, DestType := Real]" } Normalize(min := 0, value := "DiferentialPressure", max := 27648, out => "DataValues".DiferntialPressureRaw)
      { S7_Templates := "[SrcType := Real, DestType := Real]" } Scale(min := -16.0, value := "DataValues".DiferntialPressureRaw, max := 160.0, out => "DataValues".DiferntialPressure)
   END_RUNG
   // the same network as SCL:
   "DataValues".DiferntialPressureRaw := NORM_X(MIN := 0, VALUE := "DiferentialPressure", MAX := 27648);
   "DataValues".DiferntialPressure := SCALE_X(MIN := -16.0, VALUE := "DataValues".DiferntialPressureRaw, MAX := 160.0);
END_REGION

REGION Network 4: Move Differential Pressure
   RUNG wire#powerrail
      Move(in := "DataValues".DiferntialPressure, out1 => "DataValues".PipValue)
   END_RUNG
   // the same network as SCL:
   "DataValues".PipValue := "DataValues".DiferntialPressure;
END_REGION

REGION Network 5: PID REGULACION CAUDAL MOTOR
   // ENO of a box is taken as its EN; it also drops when the box reports an error
   "PID_Compact_Flow"(Setpoint := "ProcessData".PIDSetpoint,   // PID_Compact
                      Input := "ProcessData".PIDInput,
                      Input_PER := "ProcessData".PIDInput_PER,
                      ErrorAck := "ProcessData".PIDErrorAck,
                      Reset := "ProcessData".PIDReset,
                      ModeActivate := "ProcessData".PIDModeActivate,
                      Mode := "ProcessData".PIDMode,
                      Output => "ProcessData".PIDOutReal,
                      Output_PER => "ProcessData".PIDOutInt,
                      Output_PWM => "ProcessData".PIDOutPWM,
                      State => "ProcessData".PIDState,
                      Error => "ProcessData".PIDError,
                      ErrorBits => "ProcessData".PIDOutMotor);
   "ProcessData".PIDOutMotor := "ProcessData".PIDOutReal * 15.0;
END_REGION
END_ORGANIZATION_BLOCK

ORGANIZATION_BLOCK "Cyclic interrupt_PWM"   // OB31, LAD, CyclicInterrupt
{ S7_Optimized_Access := 'TRUE' }
AUTHOR : JL_Cristobal_2020
VERSION : 0.1
   VAR_INPUT
      Initial_Call : Bool;   // Initial call of this OB
      Event_Count : Int;   // Events discarded
   END_VAR
   VAR_TEMP
      Inter_Frecuency : Int;
      inter_Pulse : Int;
   END_VAR
BEGIN

REGION Network 1: Pulse Duration
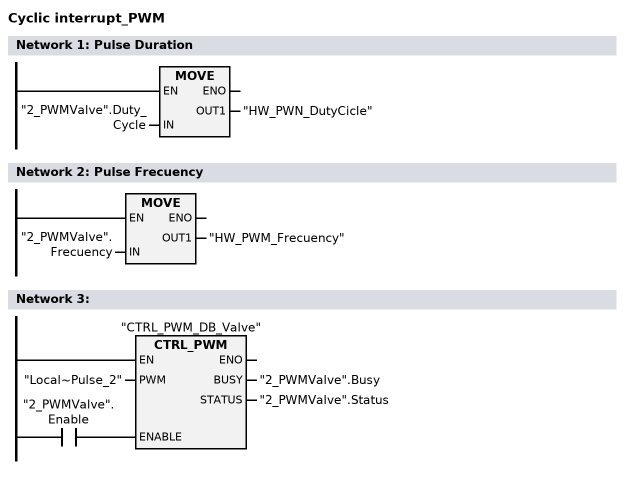
   RUNG wire#powerrail
      Move(in := "2_PWMValve".Duty_Cycle, out1 => "HW_PWN_DutyCicle")
   END_RUNG
   // the same network as SCL:
   "HW_PWN_DutyCicle" := "2_PWMValve".Duty_Cycle;
END_REGION

REGION Network 2: Pulse Frecuency
   RUNG wire#powerrail
      Move(in := "2_PWMValve".Frecuency, out1 => "HW_PWM_Frecuency")
   END_RUNG
   // the same network as SCL:
   "HW_PWM_Frecuency" := "2_PWMValve".Frecuency;
END_REGION

REGION Network 3
   "CTRL_PWM_DB_Valve"(PWM := "Local~Pulse_2",   // CTRL_PWM
                       ENABLE := "2_PWMValve".Enable,
                       BUSY => "2_PWMValve".Busy,
                       STATUS => "2_PWMValve".Status);
END_REGION
END_ORGANIZATION_BLOCK

// folder: 1_Data

FUNCTION_BLOCK "Data"   // FB10, LAD
TITLE = Data Format and Supervisor
{ S7_Optimized_Access := 'TRUE' }
AUTHOR : JL_Cristobal_2020
VERSION : 0.1
   VAR_IN_OUT
      SystemDate : Time;
      SystemTime : Time;
   END_VAR
BEGIN

REGION Network 1: Read Time and Date
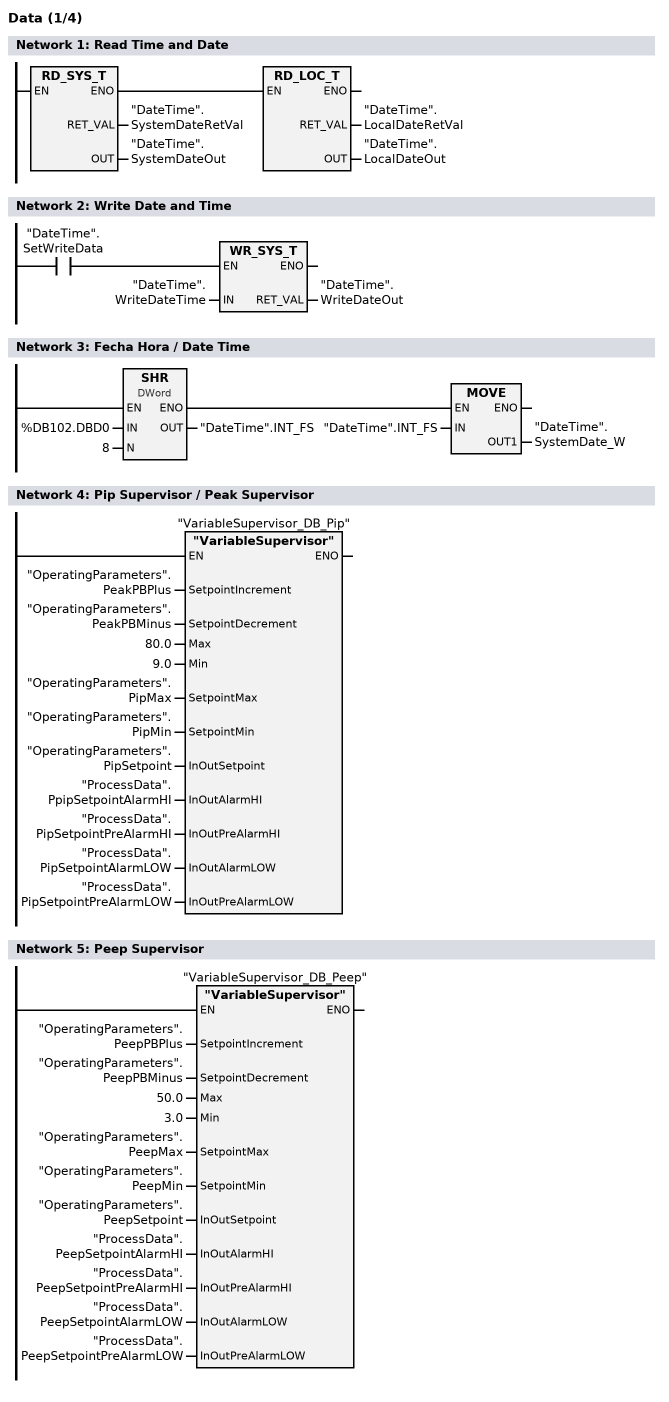
   // ENO of a box is taken as its EN; it also drops when the box reports an error
   "DateTime".SystemDateRetVal := RD_SYS_T(OUT => "DateTime".SystemDateOut);
   "DateTime".LocalDateRetVal := RD_LOC_T(OUT => "DateTime".LocalDateOut);
END_REGION

REGION Network 2: Write Date and Time
   IF "DateTime".SetWriteData THEN
       "DateTime".WriteDateOut := WR_SYS_T(IN := "DateTime".WriteDateTime);
   END_IF;
END_REGION

REGION Network 3: Fecha Hora / Date Time
   RUNG wire#powerrail
      { S7_Templates := "SrcType := DWord"; S7_GenerateENO := "TRUE" } Shr(in := %DB102.DBD0, n := 8, out => "DateTime".INT_FS)
      { S7_GenerateENO := "TRUE" } Move(in := "DateTime".INT_FS, out1 => "DateTime".SystemDate_W)
   END_RUNG
   // the same network as SCL:
   // ENO of a box is taken as its EN; it also drops when the box reports an error
   "DateTime".INT_FS := SHR(IN := %DB102.DBD0, N := 8);
   "DateTime".SystemDate_W := "DateTime".INT_FS;
END_REGION

REGION Network 4: Pip Supervisor / Peak Supervisor
   RUNG wire#powerrail
      "VariableSupervisor_DB_Pip"(SetpointIncrement := "OperatingParameters".PeakPBPlus, SetpointDecrement := "OperatingParameters".PeakPBMinus, Max := 80.0, Min := 9.0, SetpointMax := "OperatingParameters".PipMax, SetpointMin := "OperatingParameters".PipMin, InOutSetpoint := "OperatingParameters".PipSetpoint, InOutAlarmHI := "ProcessData".PpipSetpointAlarmHI, InOutPreAlarmHI := "ProcessData".PipSetpointPreAlarmHI, InOutAlarmLOW := "ProcessData".PipSetpointAlarmLOW, InOutPreAlarmLOW := "ProcessData".PipSetpointPreAlarmLOW)
   END_RUNG
   // the same network as SCL:
   "VariableSupervisor_DB_Pip"(SetpointIncrement := "OperatingParameters".PeakPBPlus,   // "VariableSupervisor"
                           SetpointDecrement := "OperatingParameters".PeakPBMinus,
                           Max := 80.0,
                           Min := 9.0,
                           SetpointMax := "OperatingParameters".PipMax,
                           SetpointMin := "OperatingParameters".PipMin,
                           InOutSetpoint := "OperatingParameters".PipSetpoint,
                           InOutAlarmHI := "ProcessData".PpipSetpointAlarmHI,
                           InOutPreAlarmHI := "ProcessData".PipSetpointPreAlarmHI,
                           InOutAlarmLOW := "ProcessData".PipSetpointAlarmLOW,
                           InOutPreAlarmLOW := "ProcessData".PipSetpointPreAlarmLOW);
END_REGION
